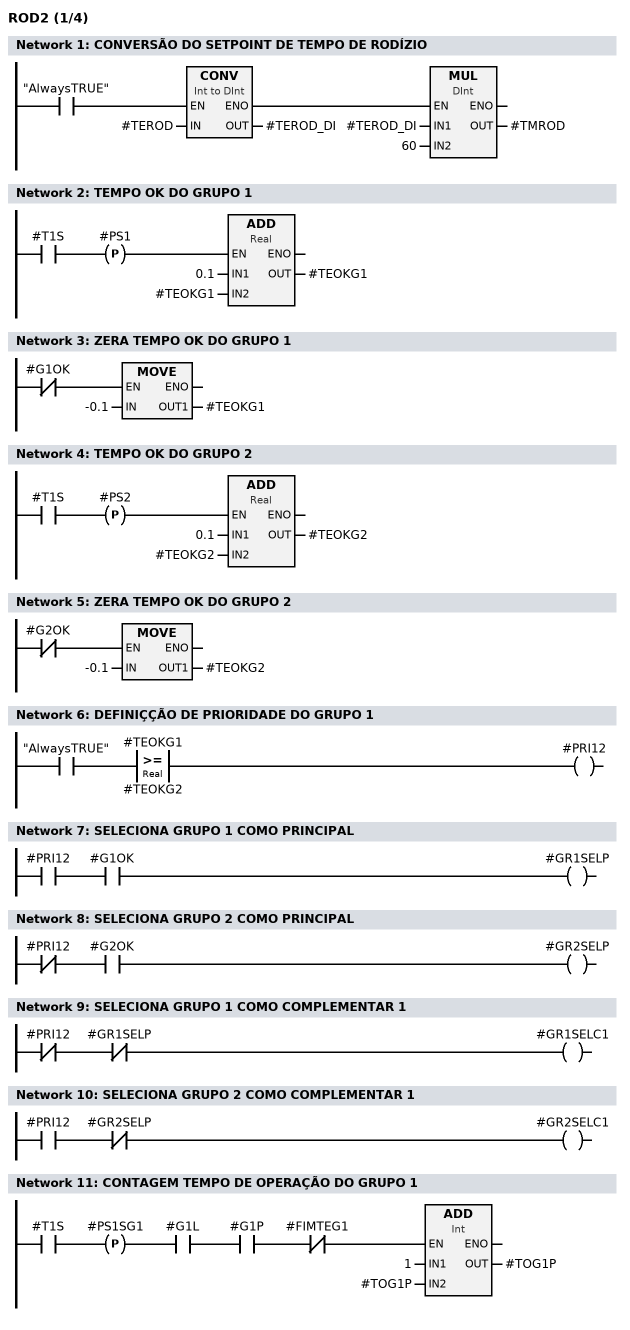
   RUNG wire#powerrail
      Contact( "AlwaysTRUE" )
      { S7_Templates := "[SrcType := Int, DestType := DInt]" } Convert(in := #TEROD, out => #TEROD_DI)
      { S7_Templates := "SrcType := DInt"; S7_GenerateENO := "TRUE" } Mul(in1 := #TEROD_DI, in2 := 60, out => #TMROD)
   END_RUNG
   // the same network as SCL:
   IF "AlwaysTRUE" THEN
       #TEROD_DI := INT_TO_DINT(#TEROD);
       #TMROD := #TEROD_DI * 60;
   END_IF;
END_REGION

REGION Network 2: TEMPO OK DO GRUPO 1
   RUNG wire#powerrail
      Contact( #T1S )
      P_Trig( #PS1 )
      { S7_Templates := "SrcType := Real"; S7_GenerateENO := "TRUE" } Add(in1 := 0.1, in2 := #TEOKG1, out => #TEOKG1)
   END_RUNG
   // the same network as SCL:
   #_w1 := #T1S AND NOT #PS1;   // rising edge
   #PS1 := #T1S;
   IF #_w1 THEN #TEOKG1 := 0.1 + #TEOKG1; END_IF;
END_REGION

REGION Network 3: ZERA TEMPO OK DO GRUPO 1
   RUNG wire#powerrail
      I_Contact( #G1OK )
      { S7_GenerateENO := "TRUE" } Move(in := -0.1, out1 => #TEOKG1)
   END_RUNG
   // the same network as SCL:
   IF NOT #G1OK THEN #TEOKG1 := -0.1; END_IF;
END_REGION

REGION Network 4: TEMPO OK DO GRUPO 2
   RUNG wire#powerrail
      Contact( #T1S )
      P_Trig( #PS2 )
      { S7_Templates := "SrcType := Real"; S7_GenerateENO := "TRUE" } Add(in1 := 0.1, in2 := #TEOKG2, out => #TEOKG2)
   END_RUNG
   // the same network as SCL:
   #_w1 := #T1S AND NOT #PS2;   // rising edge
   #PS2 := #T1S;
   IF #_w1 THEN #TEOKG2 := 0.1 + #TEOKG2; END_IF;
END_REGION

REGION Network 5: ZERA TEMPO OK DO GRUPO 2
   RUNG wire#powerrail
      I_Contact( #G2OK )
      { S7_GenerateENO := "TRUE" } Move(in := -0.1, out1 => #TEOKG2)
   END_RUNG
   // the same network as SCL:
   IF NOT #G2OK THEN #TEOKG2 := -0.1; END_IF;
END_REGION

REGION Network 6: DEFINIÇÇÃO DE PRIORIDADE DO GRUPO 1
   RUNG wire#powerrail
      Contact( "AlwaysTRUE" )
      { S7_Templates := "SrcType := Real" } GE_Contact(in1 := #TEOKG1, in2 := #TEOKG2)
      Coil( #PRI12 )
   END_RUNG
   // the same network as SCL:
   #PRI12 := "AlwaysTRUE" AND (#TEOKG1 >= #TEOKG2);
END_REGION

REGION Network 7: SELECIONA GRUPO 1 COMO PRINCIPAL
   RUNG wire#powerrail
      Contact( #PRI12 )
      Contact( #G1OK )
      Coil( #GR1SELP )
   END_RUNG
   // the same network as SCL:
   #GR1SELP := #PRI12 AND #G1OK;
END_REGION

REGION Network 8: SELECIONA GRUPO 2 COMO PRINCIPAL
   RUNG wire#powerrail
      I_Contact( #PRI12 )
      Contact( #G2OK )
      Coil( #GR2SELP )
   END_RUNG
   // the same network as SCL:
   #GR2SELP := NOT #PRI12 AND #G2OK;
END_REGION

REGION Network 9: SELECIONA GRUPO 1 COMO COMPLEMENTAR 1
   RUNG wire#powerrail
      I_Contact( #PRI12 )
      I_Contact( #GR1SELP )
      Coil( #GR1SELC1 )
   END_RUNG
   // the same network as SCL:
   #GR1SELC1 := NOT #PRI12 AND NOT #GR1SELP;
END_REGION

REGION Network 10: SELECIONA GRUPO 2 COMO COMPLEMENTAR 1
   RUNG wire#powerrail
      Contact( #PRI12 )
      I_Contact( #GR2SELP )
      Coil( #GR2SELC1 )
   END_RUNG
   // the same network as SCL:
   #GR2SELC1 := #PRI12 AND NOT #GR2SELP;
END_REGION

REGION Network 11: CONTAGEM TEMPO DE OPERAÇÃO DO GRUPO 1
   RUNG wire#powerrail
      Contact( #T1S )
      P_Trig( #PS1SG1 )
      Contact( #G1L )
      Contact( #G1P )
      I_Contact( #FIMTEG1 )
      { S7_Templates := "SrcType := Int"; S7_GenerateENO := "TRUE" } Add(in1 := 1, in2 := #TOG1P, out => #TOG1P)
   END_RUNG
   // the same network as SCL:
   #_w1 := #T1S AND NOT #PS1SG1;   // rising edge
   #PS1SG1 := #T1S;
   IF #_w1 AND #G1L AND #G1P AND NOT #FIMTEG1 THEN #TOG1P := 1 + #TOG1P; END_IF;
END_REGION

REGION Network 12: TEMPO DE OPERAÇÃO ATINGIDO
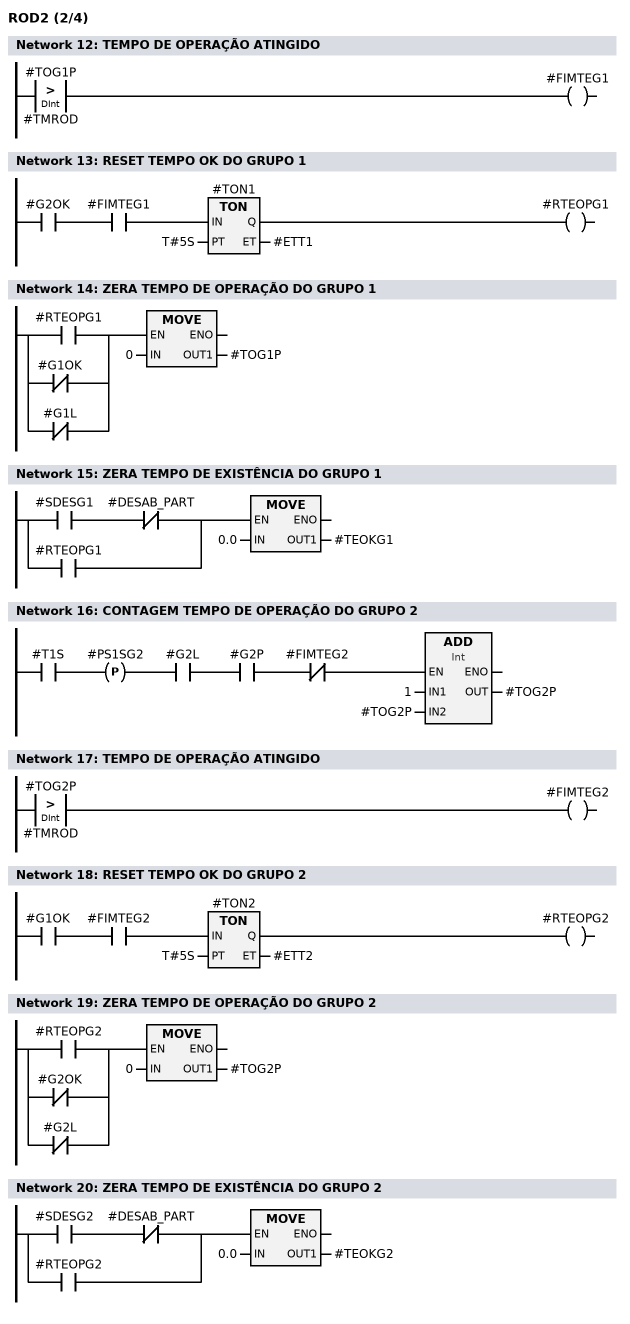
   RUNG wire#powerrail
      { S7_Templates := "SrcType := DInt" } GT_Contact(in1 := #TOG1P, in2 := #TMROD)
      Coil( #FIMTEG1 )
   END_RUNG
   // the same network as SCL:
   #FIMTEG1 := #TOG1P > #TMROD;
END_REGION

REGION Network 13: RESET TEMPO OK DO GRUPO 1
   #TON1(IN := #G2OK AND #FIMTEG1, PT := T#5S, ET => #ETT1);   // TON
   #RTEOPG1 := #TON1.Q;
END_REGION

REGION Network 14: ZERA TEMPO DE OPERAÇÃO DO GRUPO 1
   RUNG wire#powerrail
      Contact( #RTEOPG1 )
      wire#w1
      { S7_GenerateENO := "TRUE" } Move(in := 0, out1 => #TOG1P)
   END_RUNG
   RUNG wire#powerrail
      I_Contact( #G1OK )
   END_RUNG wire#w1
   RUNG wire#powerrail
      I_Contact( #G1L )
   END_RUNG wire#w1
   // the same network as SCL:
   IF #RTEOPG1 OR NOT #G1OK OR NOT #G1L THEN #TOG1P := 0; END_IF;
END_REGION

REGION Network 15: ZERA TEMPO DE EXISTÊNCIA DO GRUPO 1
   RUNG wire#powerrail
      Contact( #SDESG1 )
      I_Contact( #DESAB_PART )
      wire#w1
      { S7_GenerateENO := "TRUE" } Move(in := 0.0, out1 => #TEOKG1)
   END_RUNG
   RUNG wire#powerrail
      Contact( #RTEOPG1 )
   END_RUNG wire#w1
   // the same network as SCL:
   IF (#SDESG1 AND NOT #DESAB_PART) OR #RTEOPG1 THEN #TEOKG1 := 0.0; END_IF;
END_REGION

REGION Network 16: CONTAGEM TEMPO DE OPERAÇÃO DO GRUPO 2
   RUNG wire#powerrail
      Contact( #T1S )
      P_Trig( #PS1SG2 )
      Contact( #G2L )
      Contact( #G2P )
      I_Contact( #FIMTEG2 )
      { S7_Templates := "SrcType := Int"; S7_GenerateENO := "TRUE" } Add(in1 := 1, in2 := #TOG2P, out => #TOG2P)
   END_RUNG
   // the same network as SCL:
   #_w1 := #T1S AND NOT #PS1SG2;   // rising edge
   #PS1SG2 := #T1S;
   IF #_w1 AND #G2L AND #G2P AND NOT #FIMTEG2 THEN #TOG2P := 1 + #TOG2P; END_IF;
END_REGION

REGION Network 17: TEMPO DE OPERAÇÃO ATINGIDO
   RUNG wire#powerrail
      { S7_Templates := "SrcType := DInt" } GT_Contact(in1 := #TOG2P, in2 := #TMROD)
      Coil( #FIMTEG2 )
   END_RUNG
   // the same network as SCL:
   #FIMTEG2 := #TOG2P > #TMROD;
END_REGION

REGION Network 18: RESET TEMPO OK DO GRUPO 2
   #TON2(IN := #G1OK AND #FIMTEG2, PT := T#5S, ET => #ETT2);   // TON
   #RTEOPG2 := #TON2.Q;
END_REGION

REGION Network 19: ZERA TEMPO DE OPERAÇÃO DO GRUPO 2
   RUNG wire#powerrail
      Contact( #RTEOPG2 )
      wire#w1
      { S7_GenerateENO := "TRUE" } Move(in := 0, out1 => #TOG2P)
   END_RUNG
   RUNG wire#powerrail
      I_Contact( #G2OK )
   END_RUNG wire#w1
   RUNG wire#powerrail
      I_Contact( #G2L )
   END_RUNG wire#w1
   // the same network as SCL:
   IF #RTEOPG2 OR NOT #G2OK OR NOT #G2L THEN #TOG2P := 0; END_IF;
END_REGION

REGION Network 20: ZERA TEMPO DE EXISTÊNCIA DO GRUPO 2
   RUNG wire#powerrail
      Contact( #SDESG2 )
      I_Contact( #DESAB_PART )
      wire#w1
      { S7_GenerateENO := "TRUE" } Move(in := 0.0, out1 => #TEOKG2)
   END_RUNG
   RUNG wire#powerrail
      Contact( #RTEOPG2 )
   END_RUNG wire#w1
   // the same network as SCL:
   IF (#SDESG2 AND NOT #DESAB_PART) OR #RTEOPG2 THEN #TEOKG2 := 0.0; END_IF;
END_REGION

REGION Network 21: SELEÇÃO GRUPO 1 COMO PRINCIPAL
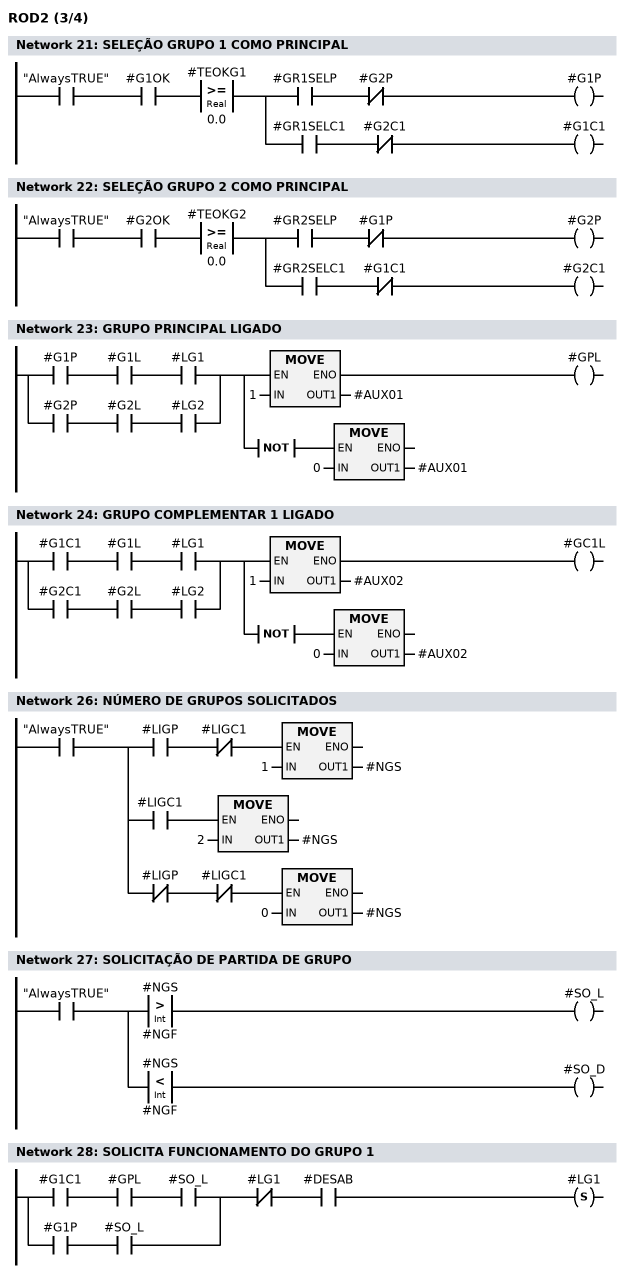
   RUNG wire#powerrail
      Contact( "AlwaysTRUE" )
      Contact( #G1OK )
      { S7_Templates := "SrcType := Real" } GE_Contact(in1 := #TEOKG1, in2 := 0.0)
      wire#w1
      Contact( #GR1SELP )
      I_Contact( #G2P )
      Coil( #G1P )
   END_RUNG
   RUNG wire#w1
      Contact( #GR1SELC1 )
      I_Contact( #G2C1 )
      Coil( #G1C1 )
   END_RUNG
   // the same network as SCL:
   #_w1 := "AlwaysTRUE" AND #G1OK AND (#TEOKG1 >= 0.0);
   #G1P := #_w1 AND #GR1SELP AND NOT #G2P;
   #G1C1 := #_w1 AND #GR1SELC1 AND NOT #G2C1;
END_REGION

REGION Network 22: SELEÇÃO GRUPO 2 COMO PRINCIPAL
   RUNG wire#powerrail
      Contact( "AlwaysTRUE" )
      Contact( #G2OK )
      { S7_Templates := "SrcType := Real" } GE_Contact(in1 := #TEOKG2, in2 := 0.0)
      wire#w1
      Contact( #GR2SELP )
      I_Contact( #G1P )
      Coil( #G2P )
   END_RUNG
   RUNG wire#w1
      Contact( #GR2SELC1 )
      I_Contact( #G1C1 )
      Coil( #G2C1 )
   END_RUNG
   // the same network as SCL:
   #_w1 := "AlwaysTRUE" AND #G2OK AND (#TEOKG2 >= 0.0);
   #G2P := #_w1 AND #GR2SELP AND NOT #G1P;
   #G2C1 := #_w1 AND #GR2SELC1 AND NOT #G1C1;
END_REGION

REGION Network 23: GRUPO PRINCIPAL LIGADO
   RUNG wire#powerrail
      Contact( #G1P )
      Contact( #G1L )
      Contact( #LG1 )
      wire#w1
      { S7_GenerateENO := "TRUE" } Move(in := 1, out1 => #AUX01)
      Coil( #GPL )
   END_RUNG
   RUNG wire#powerrail
      Contact( #G2P )
      Contact( #G2L )
      Contact( #LG2 )
   END_RUNG wire#w1
   RUNG wire#w1
      Not()
      { S7_GenerateENO := "TRUE" } Move(in := 0, out1 => #AUX01)
   END_RUNG
   // the same network as SCL:
   // ENO of a box is taken as its EN; it also drops when the box reports an error
   #_w1 := (#G1P AND #G1L AND #LG1) OR (#G2P AND #G2L AND #LG2);
   IF #_w1 THEN #AUX01 := 1; END_IF;
   #GPL := #_w1;
   IF NOT #_w1 THEN #AUX01 := 0; END_IF;
END_REGION

REGION Network 24: GRUPO COMPLEMENTAR 1 LIGADO
   RUNG wire#powerrail
      Contact( #G1C1 )
      Contact( #G1L )
      Contact( #LG1 )
      wire#w1
      { S7_GenerateENO := "TRUE" } Move(in := 1, out1 => #AUX02)
      Coil( #GC1L )
   END_RUNG
   RUNG wire#powerrail
      Contact( #G2C1 )
      Contact( #G2L )
      Contact( #LG2 )
   END_RUNG wire#w1
   RUNG wire#w1
      Not()
      { S7_GenerateENO := "TRUE" } Move(in := 0, out1 => #AUX02)
   END_RUNG
   // the same network as SCL:
   // ENO of a box is taken as its EN; it also drops when the box reports an error
   #_w1 := (#G1C1 AND #G1L AND #LG1) OR (#G2C1 AND #G2L AND #LG2);
   IF #_w1 THEN #AUX02 := 1; END_IF;
   #GC1L := #_w1;
   IF NOT #_w1 THEN #AUX02 := 0; END_IF;
END_REGION

REGION Network 25 (STL): NÚMERO DE GRUPOS FUNCIONANDO

         L     #AUX01;
         L     #AUX02;
         +I;
         T     #NGF;
END_REGION

REGION Network 26: NÚMERO DE GRUPOS SOLICITADOS
   RUNG wire#powerrail
      Contact( "AlwaysTRUE" )
      wire#w1
      Contact( #LIGP )
      I_Contact( #LIGC1 )
      { S7_GenerateENO := "TRUE" } Move(in := 1, out1 => #NGS)
   END_RUNG
   RUNG wire#w1
      Contact( #LIGC1 )
      { S7_GenerateENO := "TRUE" } Move(in := 2, out1 => #NGS)
   END_RUNG
   RUNG wire#w1
      I_Contact( #LIGP )
      I_Contact( #LIGC1 )
      { S7_GenerateENO := "TRUE" } Move(in := 0, out1 => #NGS)
   END_RUNG
   // the same network as SCL:
   IF "AlwaysTRUE" AND #LIGP AND NOT #LIGC1 THEN #NGS := 1; END_IF;
   IF "AlwaysTRUE" AND #LIGC1 THEN #NGS := 2; END_IF;
   IF "AlwaysTRUE" AND NOT #LIGP AND NOT #LIGC1 THEN #NGS := 0; END_IF;
END_REGION

REGION Network 27: SOLICITAÇÃO DE PARTIDA DE GRUPO
   RUNG wire#powerrail
      Contact( "AlwaysTRUE" )
      wire#w1
      { S7_Templates := "SrcType := Int" } GT_Contact(in1 := #NGS, in2 := #NGF)
      Coil( #SO_L )
   END_RUNG
   RUNG wire#w1
      { S7_Templates := "SrcType := Int" } LT_Contact(in1 := #NGS, in2 := #NGF)
      Coil( #SO_D )
   END_RUNG
   // the same network as SCL:
   #SO_L := "AlwaysTRUE" AND (#NGS > #NGF);
   #SO_D := "AlwaysTRUE" AND (#NGS < #NGF);
END_REGION

REGION Network 28: SOLICITA FUNCIONAMENTO DO GRUPO 1
   RUNG wire#powerrail
      Contact( #G1C1 )
      Contact( #GPL )
      Contact( #SO_L )
      wire#w1
      I_Contact( #LG1 )
      Contact( #DESAB )
      S_Coil( #LG1 )
   END_RUNG
   RUNG wire#powerrail
      Contact( #G1P )
      Contact( #SO_L )
   END_RUNG wire#w1
   // the same network as SCL:
   IF ((#G1C1 AND #GPL AND #SO_L) OR (#G1P AND #SO_L)) AND NOT #LG1 AND #DESAB THEN #LG1 := TRUE; END_IF;
END_REGION

REGION Network 29: SOLICITA FUNCIONAMENTO DO GRUPO 2
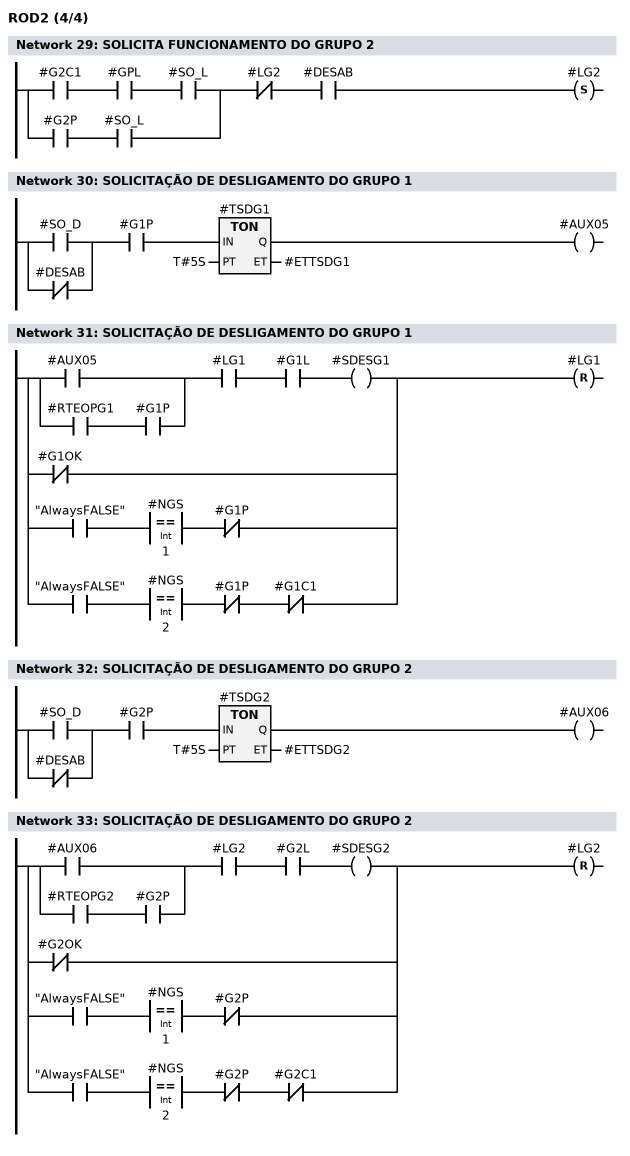
   RUNG wire#powerrail
      Contact( #G2C1 )
      Contact( #GPL )
      Contact( #SO_L )
      wire#w1
      I_Contact( #LG2 )
      Contact( #DESAB )
      S_Coil( #LG2 )
   END_RUNG
   RUNG wire#powerrail
      Contact( #G2P )
      Contact( #SO_L )
   END_RUNG wire#w1
   // the same network as SCL:
   IF ((#G2C1 AND #GPL AND #SO_L) OR (#G2P AND #SO_L)) AND NOT #LG2 AND #DESAB THEN #LG2 := TRUE; END_IF;
END_REGION

REGION Network 30: SOLICITAÇÃO DE DESLIGAMENTO DO GRUPO 1
   #TSDG1(IN := (#SO_D OR NOT #DESAB) AND #G1P, PT := T#5S, ET => #ETTSDG1);   // TON
   #AUX05 := #TSDG1.Q;
END_REGION

REGION Network 31: SOLICITAÇÃO DE DESLIGAMENTO DO GRUPO 1
   RUNG wire#powerrail
      Contact( #AUX05 )
      wire#w1
      Contact( #LG1 )
      Contact( #G1L )
      Coil( #SDESG1 )
      wire#w2
      R_Coil( #LG1 )
   END_RUNG
   RUNG wire#powerrail
      Contact( #RTEOPG1 )
      Contact( #G1P )
   END_RUNG wire#w1
   RUNG wire#powerrail
      I_Contact( #G1OK )
   END_RUNG wire#w2
   RUNG wire#powerrail
      Contact( "AlwaysFALSE" )
      { S7_Templates := "SrcType := Int" } EQ_Contact(in1 := #NGS, in2 := 1)
      I_Contact( #G1P )
   END_RUNG wire#w2
   RUNG wire#powerrail
      Contact( "AlwaysFALSE" )
      { S7_Templates := "SrcType := Int" } EQ_Contact(in1 := #NGS, in2 := 2)
      I_Contact( #G1P )
      I_Contact( #G1C1 )
   END_RUNG wire#w2
   // the same network as SCL:
   #SDESG1 := (#AUX05 OR (#RTEOPG1 AND #G1P)) AND #LG1 AND #G1L;
   IF #SDESG1 OR NOT #G1OK OR ("AlwaysFALSE" AND (#NGS = 1) AND NOT #G1P) OR ("AlwaysFALSE" AND (#NGS = 2) AND NOT #G1P AND NOT #G1C1) THEN
       #LG1 := FALSE;
   END_IF;
END_REGION

REGION Network 32: SOLICITAÇÃO DE DESLIGAMENTO DO GRUPO 2
   #TSDG2(IN := (#SO_D OR NOT #DESAB) AND #G2P, PT := T#5S, ET => #ETTSDG2);   // TON
   #AUX06 := #TSDG2.Q;
END_REGION

REGION Network 33: SOLICITAÇÃO DE DESLIGAMENTO DO GRUPO 2
   RUNG wire#powerrail
      Contact( #AUX06 )
      wire#w1
      Contact( #LG2 )
      Contact( #G2L )
      Coil( #SDESG2 )
      wire#w2
      R_Coil( #LG2 )
   END_RUNG
   RUNG wire#powerrail
      Contact( #RTEOPG2 )
      Contact( #G2P )
   END_RUNG wire#w1
   RUNG wire#powerrail
      I_Contact( #G2OK )
   END_RUNG wire#w2
   RUNG wire#powerrail
      Contact( "AlwaysFALSE" )
      { S7_Templates := "SrcType := Int" } EQ_Contact(in1 := #NGS, in2 := 1)
      I_Contact( #G2P )
   END_RUNG wire#w2
   RUNG wire#powerrail
      Contact( "AlwaysFALSE" )
      { S7_Templates := "SrcType := Int" } EQ_Contact(in1 := #NGS, in2 := 2)
      I_Contact( #G2P )
      I_Contact( #G2C1 )
   END_RUNG wire#w2
   // the same network as SCL:
   #SDESG2 := (#AUX06 OR (#RTEOPG2 AND #G2P)) AND #LG2 AND #G2L;
   IF #SDESG2 OR NOT #G2OK OR ("AlwaysFALSE" AND (#NGS = 1) AND NOT #G2P) OR ("AlwaysFALSE" AND (#NGS = 2) AND NOT #G2P AND NOT #G2C1) THEN
       #LG2 := FALSE;
   END_IF;
END_REGION
END_FUNCTION_BLOCK

FUNCTION_BLOCK "DANFOSS_REV"   // FB206, LAD
TITLE = CONTROLE INVERSOR SINAMICS
{ S7_Optimized_Access := 'FALSE' }
VERSION : 0.1
   VAR_INPUT
      DBNO : Int;   // Número do DB
      DBPOS : Int;   // Posição do DB
      MF1 : Bool;   // Motor em falha
      MF2 : Bool;   // Motor em falha
      HM : Bool;   // Habilita manual
      HA : Bool;   // Habilita automático
      HAR : Bool;   // Habilita automático reverso
      CMA : Bool;   // Comando liga automático
      CLM : Bool;   // Comando liga manual
      CLMR : Bool;   // Comando liga manual reverso
      CDM : Bool;   // Comando desliga manual
      CRF : Bool;   // Comando reset de falha
      CRTO : Bool;   // Comando reset tepo de operação
      CHC : Bool;   // Comando habilita controle de velocidade
      CHB : Bool;   // Comando habilita bloqueio
      CL1S : Bool;   // Pulso a cada 1 segundo
      SRC : Bool;   // Status rede de comunicação
      FMM : Real;   // Fundo de escala frequência do motor
      SPM : Real;   // Setpoint manual de velocidade
      SPA : Real;   // Setpoint automático de velocidade
   END_VAR
   VAR_OUTPUT
      YFL : Bool;   // Indicação de falha no inversor
      YFPP : Bool;   // Indicação de falha no acionamento
      YR : Bool;   // Indicação de chave na posição remota
      YSH : Bool;   // Indicação de motor ligado
      YF : Bool;   // Indicação de motor em falha
      CL : Bool;   // Comando liga motor
      REV : Bool;   // Indicação de motor ligado no sentido reverso
      CMD_RESET : Bool;   // Reset de falha
      IN18 : Bool;   // ENTRADA DIGITAL
      IN19 : Bool;   // ENTRADA DIGITAL
      IN27 : Bool;   // ENTRADA DIGITAL
      IN29 : Bool;   // ENTRADA DIGITAL
      IN32 : Bool;   // ENTRADA DIGITAL
      IN33 : Bool;   // ENTRADA DIGITAL
      IT : Real;   // Indicação de corrente
      ST : Real;   // Indicação de frequência
   END_VAR
   VAR_IN_OUT
      SEG : Int;   // Segundos de operação
      MIN : Int;   // Minutos de operação
      HOR : Int;   // Horas de operação
   END_VAR
   VAR
      STW : Struct   // PALAVRA DE STATUS DO INVERSOR
         SpeddRef : Bool;   // Velocidade=Setpoint
         BUS : Bool;   // Controle pelo BUS
         FreqOK : Bool;   // Frequecia OK
         Operation : Bool;   // Em operação
         Drive : Bool;   // Drive OK
         Voltage : Bool;   // Tensão excedida
         Torque : Bool;   // Torque excedido
         Thermal : Bool;   // Térmico excedido
         Ready_forswitch_on : Bool;   // Controle habilitado
         Ready : Bool;   // Inversor pronto
         Running : Bool;   // Em funcionamento
         Fault : Bool;   // Falha ativa
         Error : Bool;   // Erro ativo
         Reservado : Bool;   // Reservado
         TripLock : Bool;   // Inibição ativa
         Warning : Bool;   // Advertência
      END_STRUCT;
      LPZD2 : Int;   // Velocidade do motor
      LPZD3 : Int;   // Corrente do motor
      LPZD4 : Struct   // Entradas digitais
         INX2 : Bool;   // Reservado
         INX3 : Bool;   // Reservado
         INX4 : Bool;   // Reservado
         INX5 : Bool;   // Reservado
         INX6 : Bool;   // Reservado
         INX7 : Bool;   // Reservado
         INX8 : Bool;   // Reservado
         INX9 : Bool;   // Reservado
         IN33 : Bool;   // Entrada terminal 33
         IN32 : Bool;   // Entrada terminal 32
         IN29 : Bool;   // Entrada terminal 29
         IN27 : Bool;   // Entrada terminal 27
         IN19 : Bool;   // Entrada terminal 19
         IN18 : Bool;   // Entrada terminal 18
         INX0 : Bool;   // Reservado
         INX1 : Bool;   // Reservado
      END_STRUCT;
      CTW : Struct   // PALAVRA DE CONTROLE DO INVERSOR
         Jog : Bool;   // Habilita jog
         RampSEL : Bool;   // Seleção RAMPA1/2
         Control_plc : Bool;   // Valida dados do PLC
         Relay1 : Bool;   // Habilita partida sentido reverso
         Relay4 : Bool;   // Controlador de velocidade habilitado
         Setup0 : Bool;   // Seleção de setup bit0
         Setup1 : Bool;   // Seleção de setup bit1
         Start_reverse : Bool;   // Habilita partida sentido reverso
         LSB : Bool;   // Seleção externa LSB
         MSB : Bool;   // Seleção externa MSB
         DCbrakeRamp : Bool;   // Freio DC/Rampa
         Coasting : Bool;   // Liga motor
         Enable_Ramp : Bool;   // Habilita rampa
         Enable_ramp_generator : Bool;   // Habilita gerador de rampa
         Start : Bool;   // Liga motor
         Reset : Bool;   // Reconhecimento de falha
      END_STRUCT;
      CT_MotorReference : Int;   // Referência de velocidade
      EPZD3 : Int;   // Reserva
      EPZD4 : Int;   // Reserva
      RESET : Bool;   // Reset de falha
      AUX01 : Bool;   // Auxiliar utilizado na lógica
      AUX02 : Bool;   // Auxiliar utilizado na lógica
      AUX03 : Bool;   // Auxiliar utilizado na lógica
      AUX04 : Bool;   // Auxiliar utilizado na lógica
      AUX05 : Bool;   // Auxiliar utilizado na lógica
      AUX06 : Bool;   // Auxiliar utilizado na lógica
      AUX07 : Bool;   // Auxiliar utilizado na lógica
      AUX08 : Bool;   // Auxiliar utilizado na lógica
      AUX09 : Bool;   // Auxiliar utilizado na lógica
      AUX10 : Bool;   // Auxiliar utilizado na lógica
      P60S : Bool;   // Pulso de 60 segundos
      P60M : Bool;   // Pulso de 60 minutos
      PFHO : Bool;   // Pulso de limite de horas
      SPS : Real;   // Frequência para controle
      TPP1 : TON_TIME;   // Temporizador falha no acionamento
      TPP2 : TON_TIME;   // Temporizador falha no acionamento
      TR : TON_TIME;   // Temporizador reset de falha
   END_VAR
   VAR_TEMP
      LIGADO : Bool;   // Ligado
      FALHA : Bool;   // Falha
      TEMP0 : Bool;
      TEMP1 : Bool;
      ET_TPP1 : Time;   // Efetivo temporizador
      ET_TPP2 : Time;   // Efetivo temporizador
      ET_TR : Time;   // Efetivo temporizador
      AUXDB : Int;   // Auxiliar movimentação do DB
      ST1 : Real;   // Frequência convertida
   END_VAR
   VAR_TEMP   // added for the SCL form of the ladder/FBD networks
      _w1 : Bool;
      _w2 : Bool;
      _w3 : Bool;
      _w4 : Bool;
   END_VAR
BEGIN

REGION Network 1 (STL): Leitura de dados da rede
   //CARREGA O ENDEREÇO DA PRIMEIRA WORD DE ENTRADA

         L     #DBNO;  // Carrega n° da DB
         T     #AUXDB;

         OPN   DB[ #AUXDB];  // Abre DB

         L     #DBPOS;  // Multiplica valor da posição para acertar ponteiro (valor x 8bit´s)
         L     8;
         *I;
         LAR1;  // Carrega valor de ponteiro no registrador 1

         L     DBW [ AR1 , P#0.0 ];
         T     %XDataW34;
         L     DBW [ AR1 , P#2.0 ];
         T     #LPZD2;
         L     DBW [ AR1 , P#4.0 ];
         T     #LPZD3;
         L     DBW [ AR1 , P#6.0 ];
         T     %XDataW40;
END_REGION

REGION Network 2 (STL): CONVERSÃO DA LEITURA DE FREQUÊNCIA/CORRENTE
         L     #LPZD2;
         ITD;
         DTR;
         L     #FMM;
         *R;
         L     16384.0;
         /R;
         T     #ST;

         L     #LPZD3;
         ITD;
         DTR;
         L     100.0;
         /R;
         T     #IT;
END_REGION

REGION Network 3 (STL): STATUS DO INVERSOR
   // VERIFICA ESTADO DO PRIMEIRO BYTE DA PALAVRA DE ENTRADA  (PZD)

         A     #STW.Fault;
         =     #YFL;  //ALARME DE FALHA NO INVERSOR

   // LEITURA DAS ENTRADAS DIGITAIS

         A     #LPZD4.IN33;  // ENTRADA DIGITAL DE REMOTO
         A     #STW.BUS;
         =     #YR;
         =     #IN33;

         A     #LPZD4.IN18;  // TERMINAL 18
         =     #IN18;

         A     #LPZD4.IN19;  // TERMINAL 19
         =     #IN19;

         A     #LPZD4.IN27;  // TERMINAL 27
         =     #IN27;

         A     #LPZD4.IN32;  // TERMINAL 32
         =     #IN32;

         A     #LPZD4.IN29;  // TERMINAL 29
         =     #IN29;
END_REGION

REGION Network 4: STATUS DE LIGADO
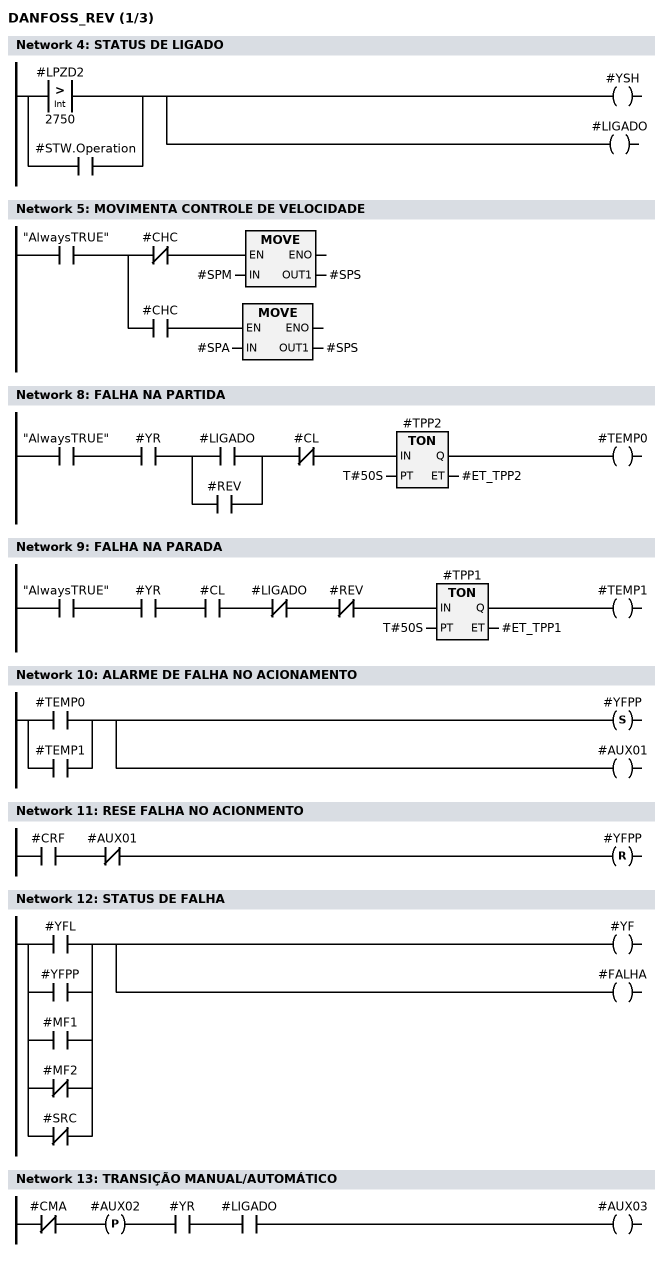
   RUNG wire#powerrail
      { S7_Templates := "SrcType := Int" } GT_Contact(in1 := #LPZD2, in2 := 2750)
      wire#w1
      Coil( #YSH )
   END_RUNG
   RUNG wire#powerrail
      Contact( #STW.Operation )
   END_RUNG wire#w1
   RUNG wire#w1
      Coil( #LIGADO )
   END_RUNG
   // the same network as SCL:
   #YSH := (#LPZD2 > 2750) OR #STW.Operation;
   #LIGADO := #YSH;
END_REGION

REGION Network 5: MOVIMENTA CONTROLE DE VELOCIDADE
   RUNG wire#powerrail
      Contact( "AlwaysTRUE" )
      wire#w1
      I_Contact( #CHC )
      { S7_GenerateENO := "TRUE" } Move(in := #SPM, out1 => #SPS)
   END_RUNG
   RUNG wire#w1
      Contact( #CHC )
      { S7_GenerateENO := "TRUE" } Move(in := #SPA, out1 => #SPS)
   END_RUNG
   // the same network as SCL:
   IF "AlwaysTRUE" AND NOT #CHC THEN #SPS := #SPM; END_IF;
   IF "AlwaysTRUE" AND #CHC THEN #SPS := #SPA; END_IF;
END_REGION

REGION Network 6 (STL): Escreve setpoint de velocidade no inversor
         L     16384.0;  //Divide para encontrar a relação de conversão
         L     #SPS;
         *R;

         L     #FMM;  //Multiplica setpoint por fator para envio ao inversor
         /R;
         RND;
         T     #CT_MotorReference;
END_REGION

REGION Network 7 (STL): ESCRITA DE DADOS NO INVERSOR
         +AR1  P#20.0;  //Carrega posição de escrita da DB

         L     %XDataW42;
         T     DBW [ AR1 , P#0.0 ];  //Offset inicial
         L     #CT_MotorReference;
         T     DBW [ AR1 , P#2.0 ];
END_REGION

REGION Network 8: FALHA NA PARTIDA
   #TPP2(IN := "AlwaysTRUE" AND #YR AND (#LIGADO OR #REV) AND NOT #CL, PT := T#50S, ET => #ET_TPP2);   // TON
   #TEMP0 := #TPP2.Q;
END_REGION

REGION Network 9: FALHA NA PARADA
   #TPP1(IN := "AlwaysTRUE" AND #YR AND #CL AND NOT #LIGADO AND NOT #REV, PT := T#50S, ET => #ET_TPP1);   // TON
   #TEMP1 := #TPP1.Q;
END_REGION

REGION Network 10: ALARME DE FALHA NO ACIONAMENTO
   RUNG wire#powerrail
      Contact( #TEMP0 )
      wire#w1
      S_Coil( #YFPP )
   END_RUNG
   RUNG wire#powerrail
      Contact( #TEMP1 )
   END_RUNG wire#w1
   RUNG wire#w1
      Coil( #AUX01 )
   END_RUNG
   // the same network as SCL:
   #_w1 := #TEMP0 OR #TEMP1;
   IF #_w1 THEN #YFPP := TRUE; END_IF;
   #AUX01 := #_w1;
END_REGION

REGION Network 11: RESE FALHA NO ACIONMENTO
   RUNG wire#powerrail
      Contact( #CRF )
      I_Contact( #AUX01 )
      R_Coil( #YFPP )
   END_RUNG
   // the same network as SCL:
   IF #CRF AND NOT #AUX01 THEN #YFPP := FALSE; END_IF;
END_REGION

REGION Network 12: STATUS DE FALHA
   RUNG wire#powerrail
      Contact( #YFL )
      wire#w1
      Coil( #YF )
   END_RUNG
   RUNG wire#powerrail
      Contact( #YFPP )
   END_RUNG wire#w1
   RUNG wire#powerrail
      Contact( #MF1 )
   END_RUNG wire#w1
   RUNG wire#powerrail
      I_Contact( #MF2 )
   END_RUNG wire#w1
   RUNG wire#powerrail
      I_Contact( #SRC )
   END_RUNG wire#w1
   RUNG wire#w1
      Coil( #FALHA )
   END_RUNG
   // the same network as SCL:
   #YF := #YFL OR #YFPP OR #MF1 OR NOT #MF2 OR NOT #SRC;
   #FALHA := #YF;
END_REGION

REGION Network 13: TRANSIÇÃO MANUAL/AUTOMÁTICO
   RUNG wire#powerrail
      I_Contact( #CMA )
      P_Trig( #AUX02 )
      Contact( #YR )
      Contact( #LIGADO )
      Coil( #AUX03 )
   END_RUNG
   // the same network as SCL:
   #_w1 := NOT #CMA AND NOT #AUX02;   // rising edge
   #AUX02 := NOT #CMA;
   #AUX03 := #_w1 AND #YR AND #LIGADO;
END_REGION

REGION Network 14: COMANDO LIGA MANUAL SENTIDO DIRETO
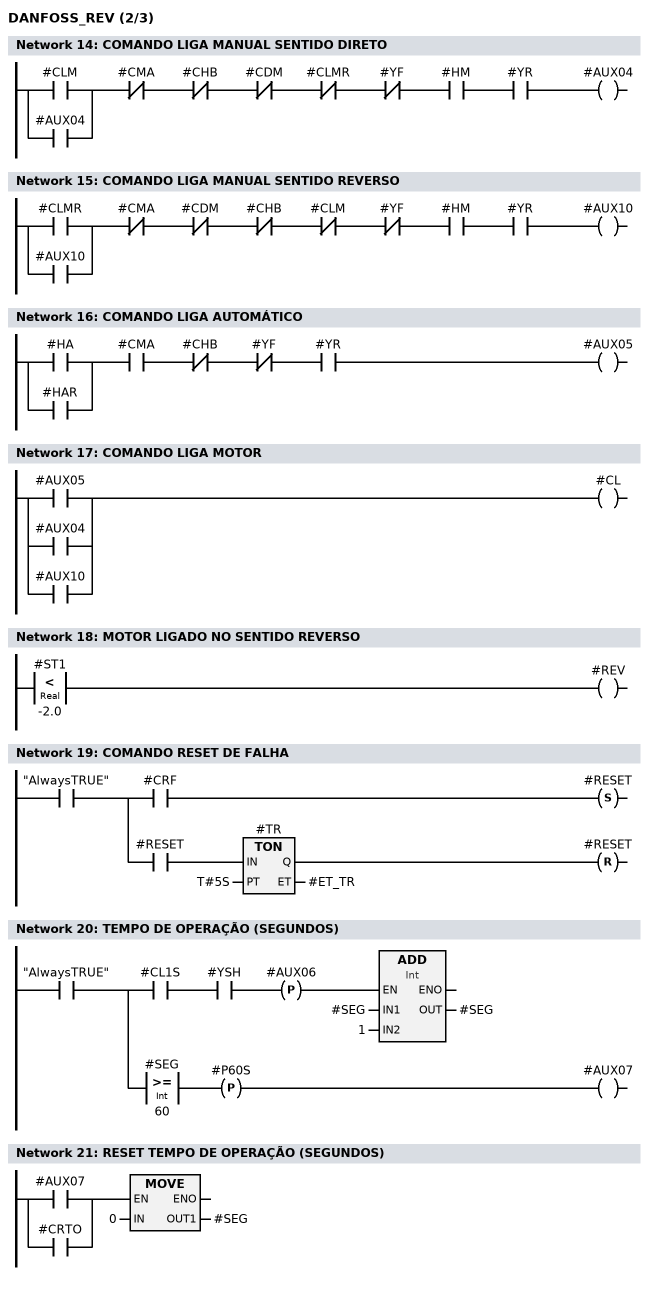
   RUNG wire#powerrail
      Contact( #CLM )
      wire#w1
      I_Contact( #CMA )
      I_Contact( #CHB )
      I_Contact( #CDM )
      I_Contact( #CLMR )
      I_Contact( #YF )
      Contact( #HM )
      Contact( #YR )
      Coil( #AUX04 )
   END_RUNG
   RUNG wire#powerrail
      Contact( #AUX04 )
   END_RUNG wire#w1
   // the same network as SCL:
   #AUX04 := (#CLM OR #AUX04) AND NOT #CMA AND NOT #CHB AND NOT #CDM AND NOT #CLMR AND NOT #YF AND #HM AND #YR;
END_REGION

REGION Network 15: COMANDO LIGA MANUAL SENTIDO REVERSO
   RUNG wire#powerrail
      Contact( #CLMR )
      wire#w1
      I_Contact( #CMA )
      I_Contact( #CDM )
      I_Contact( #CHB )
      I_Contact( #CLM )
      I_Contact( #YF )
      Contact( #HM )
      Contact( #YR )
      Coil( #AUX10 )
   END_RUNG
   RUNG wire#powerrail
      Contact( #AUX10 )
   END_RUNG wire#w1
   // the same network as SCL:
   #AUX10 := (#CLMR OR #AUX10) AND NOT #CMA AND NOT #CDM AND NOT #CHB AND NOT #CLM AND NOT #YF AND #HM AND #YR;
END_REGION

REGION Network 16: COMANDO LIGA AUTOMÁTICO
   RUNG wire#powerrail
      Contact( #HA )
      wire#w1
      Contact( #CMA )
      I_Contact( #CHB )
      I_Contact( #YF )
      Contact( #YR )
      Coil( #AUX05 )
   END_RUNG
   RUNG wire#powerrail
      Contact( #HAR )
   END_RUNG wire#w1
   // the same network as SCL:
   #AUX05 := (#HA OR #HAR) AND #CMA AND NOT #CHB AND NOT #YF AND #YR;
END_REGION

REGION Network 17: COMANDO LIGA MOTOR
   RUNG wire#powerrail
      Contact( #AUX05 )
      wire#w1
      Coil( #CL )
   END_RUNG
   RUNG wire#powerrail
      Contact( #AUX04 )
   END_RUNG wire#w1
   RUNG wire#powerrail
      Contact( #AUX10 )
   END_RUNG wire#w1
   // the same network as SCL:
   #CL := #AUX05 OR #AUX04 OR #AUX10;
END_REGION

REGION Network 18: MOTOR LIGADO NO SENTIDO REVERSO
   RUNG wire#powerrail
      { S7_Templates := "SrcType := Real" } LT_Contact(in1 := #ST1, in2 := -2.0)
      Coil( #REV )
   END_RUNG
   // the same network as SCL:
   #REV := #ST1 < (-2.0);
END_REGION

REGION Network 19: COMANDO RESET DE FALHA
   IF "AlwaysTRUE" AND #CRF THEN #RESET := TRUE; END_IF;
   #TR(IN := "AlwaysTRUE" AND #RESET, PT := T#5S, ET => #ET_TR);   // TON
   IF #TR.Q THEN #RESET := FALSE; END_IF;
END_REGION

REGION Network 20: TEMPO DE OPERAÇÃO (SEGUNDOS)
   RUNG wire#powerrail
      Contact( "AlwaysTRUE" )
      wire#w1
      Contact( #CL1S )
      Contact( #YSH )
      P_Trig( #AUX06 )
      { S7_Templates := "SrcType := Int"; S7_GenerateENO := "TRUE" } Add(in1 := #SEG, in2 := 1, out => #SEG)
   END_RUNG
   RUNG wire#w1
      { S7_Templates := "SrcType := Int" } GE_Contact(in1 := #SEG, in2 := 60)
      P_Trig( #P60S )
      Coil( #AUX07 )
   END_RUNG
   // the same network as SCL:
   #_w1 := "AlwaysTRUE" AND #CL1S AND #YSH;
   #_w2 := #_w1 AND NOT #AUX06;   // rising edge
   #AUX06 := #_w1;
   IF #_w2 THEN #SEG := #SEG + 1; END_IF;
   #_w3 := "AlwaysTRUE" AND (#SEG >= 60);
   #_w4 := #_w3 AND NOT #P60S;   // rising edge
   #P60S := #_w3;
   #AUX07 := #_w4;
END_REGION

REGION Network 21: RESET TEMPO DE OPERAÇÃO (SEGUNDOS)
   RUNG wire#powerrail
      Contact( #AUX07 )
      wire#w1
      { S7_GenerateENO := "TRUE" } Move(in := 0, out1 => #SEG)
   END_RUNG
   RUNG wire#powerrail
      Contact( #CRTO )
   END_RUNG wire#w1
   // the same network as SCL:
   IF #AUX07 OR #CRTO THEN #SEG := 0; END_IF;
END_REGION

REGION Network 22: TEMPO DE OPERAÇÃO (MINUTOS)
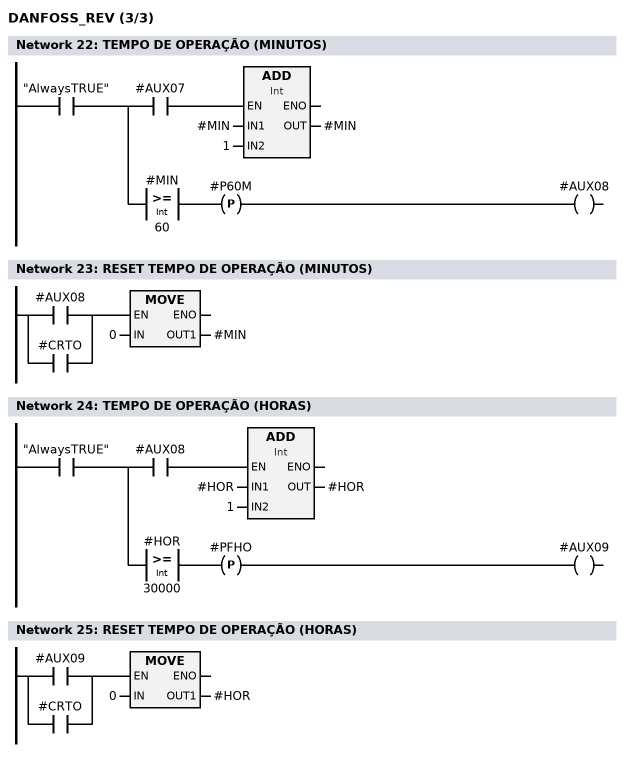
   RUNG wire#powerrail
      Contact( "AlwaysTRUE" )
      wire#w1
      Contact( #AUX07 )
      { S7_Templates := "SrcType := Int"; S7_GenerateENO := "TRUE" } Add(in1 := #MIN, in2 := 1, out => #MIN)
   END_RUNG
   RUNG wire#w1
      { S7_Templates := "SrcType := Int" } GE_Contact(in1 := #MIN, in2 := 60)
      P_Trig( #P60M )
      Coil( #AUX08 )
   END_RUNG
   // the same network as SCL:
   IF "AlwaysTRUE" AND #AUX07 THEN #MIN := #MIN + 1; END_IF;
   #_w1 := "AlwaysTRUE" AND (#MIN >= 60);
   #_w2 := #_w1 AND NOT #P60M;   // rising edge
   #P60M := #_w1;
   #AUX08 := #_w2;
END_REGION

REGION Network 23: RESET TEMPO DE OPERAÇÃO (MINUTOS)
   RUNG wire#powerrail
      Contact( #AUX08 )
      wire#w1
      { S7_GenerateENO := "TRUE" } Move(in := 0, out1 => #MIN)
   END_RUNG
   RUNG wire#powerrail
      Contact( #CRTO )
   END_RUNG wire#w1
   // the same network as SCL:
   IF #AUX08 OR #CRTO THEN #MIN := 0; END_IF;
END_REGION

REGION Network 24: TEMPO DE OPERAÇÃO (HORAS)
   RUNG wire#powerrail
      Contact( "AlwaysTRUE" )
      wire#w1
      Contact( #AUX08 )
      { S7_Templates := "SrcType := Int"; S7_GenerateENO := "TRUE" } Add(in1 := #HOR, in2 := 1, out => #HOR)
   END_RUNG
   RUNG wire#w1
      { S7_Templates := "SrcType := Int" } GE_Contact(in1 := #HOR, in2 := 30000)
      P_Trig( #PFHO )
      Coil( #AUX09 )
   END_RUNG
   // the same network as SCL:
   IF "AlwaysTRUE" AND #AUX08 THEN #HOR := #HOR + 1; END_IF;
   #_w1 := "AlwaysTRUE" AND (#HOR >= 30000);
   #_w2 := #_w1 AND NOT #PFHO;   // rising edge
   #PFHO := #_w1;
   #AUX09 := #_w2;
END_REGION
